REGION Network 156
   RUNG wire#powerrail
      Move(in := "Carrier_57_SDCFaultCode", out1 => "DB_SDC_EMS_TA".EMS[57].TA[1].FAULT)
      wire#w1
      Move(in := "Carrier_57_SDCFaultCode", out1 => "EMS".Carrier[57].SDC_IN.CarrierDriveFaults)
   END_RUNG
   RUNG wire#powerrail
      Contact( "IndiconTempDebugON" )
   END_RUNG wire#w1
   // the same network as SCL:
   "DB_SDC_EMS_TA".EMS[57].TA[1].FAULT := "Carrier_57_SDCFaultCode";
   IF TRUE OR "IndiconTempDebugON" THEN
       "EMS".Carrier[57].SDC_IN.CarrierDriveFaults := "Carrier_57_SDCFaultCode";
   END_IF;
END_REGION

REGION Network 157
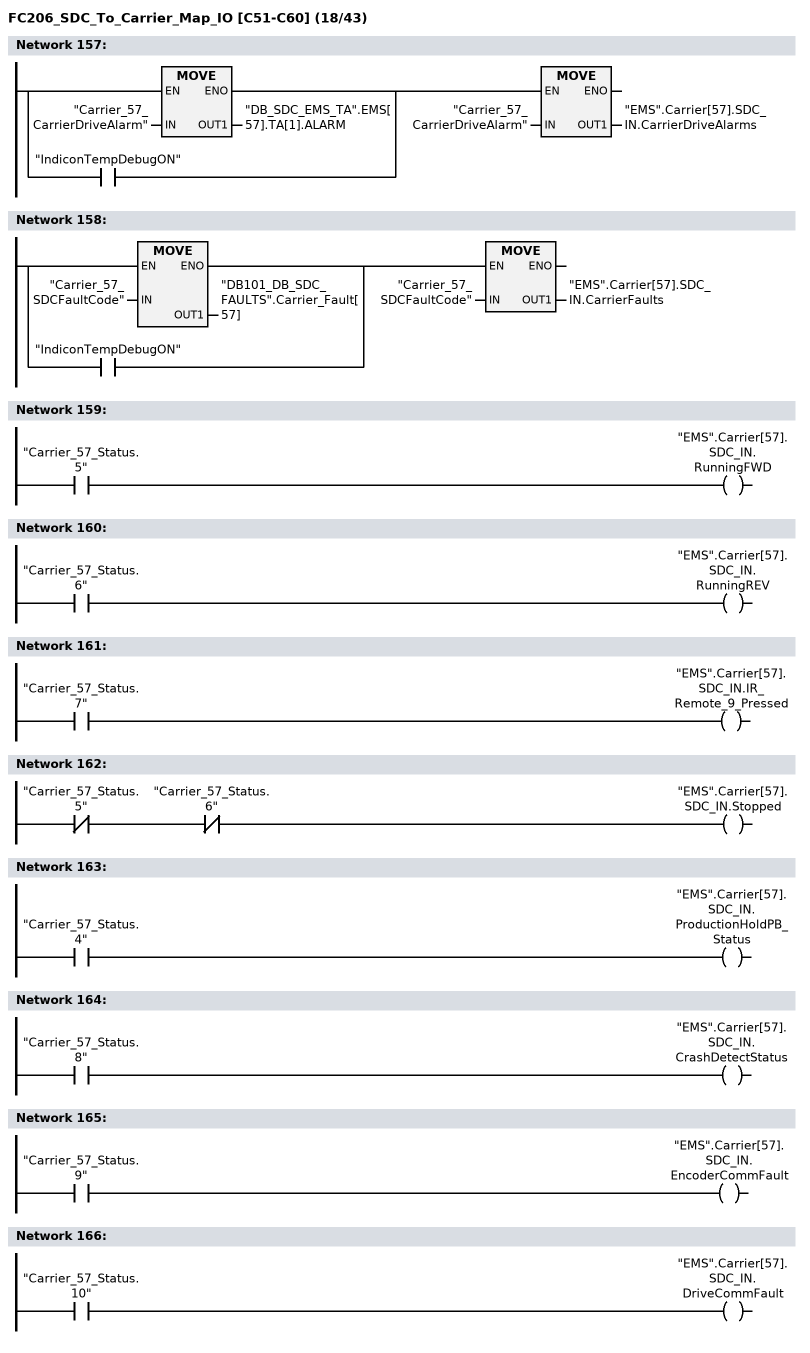
   RUNG wire#powerrail
      Move(in := "Carrier_57_CarrierDriveAlarm", out1 => "DB_SDC_EMS_TA".EMS[57].TA[1].ALARM)
      wire#w1
      Move(in := "Carrier_57_CarrierDriveAlarm", out1 => "EMS".Carrier[57].SDC_IN.CarrierDriveAlarms)
   END_RUNG
   RUNG wire#powerrail
      Contact( "IndiconTempDebugON" )
   END_RUNG wire#w1
   // the same network as SCL:
   "DB_SDC_EMS_TA".EMS[57].TA[1].ALARM := "Carrier_57_CarrierDriveAlarm";
   IF TRUE OR "IndiconTempDebugON" THEN
       "EMS".Carrier[57].SDC_IN.CarrierDriveAlarms := "Carrier_57_CarrierDriveAlarm";
   END_IF;
END_REGION

REGION Network 158
   RUNG wire#powerrail
      Move(in := "Carrier_57_SDCFaultCode", out1 => "DB101_DB_SDC_FAULTS".Carrier_Fault[57])
      wire#w1
      Move(in := "Carrier_57_SDCFaultCode", out1 => "EMS".Carrier[57].SDC_IN.CarrierFaults)
   END_RUNG
   RUNG wire#powerrail
      Contact( "IndiconTempDebugON" )
   END_RUNG wire#w1
   // the same network as SCL:
   "DB101_DB_SDC_FAULTS".Carrier_Fault[57] := "Carrier_57_SDCFaultCode";
   IF TRUE OR "IndiconTempDebugON" THEN
       "EMS".Carrier[57].SDC_IN.CarrierFaults := "Carrier_57_SDCFaultCode";
   END_IF;
END_REGION

REGION Network 159
   RUNG wire#powerrail
      Contact( "Carrier_57_Status.5" )
      Coil( "EMS".Carrier[57].SDC_IN.RunningFWD )
   END_RUNG
   // the same network as SCL:
   "EMS".Carrier[57].SDC_IN.RunningFWD := "Carrier_57_Status.5";
END_REGION

REGION Network 160
   RUNG wire#powerrail
      Contact( "Carrier_57_Status.6" )
      Coil( "EMS".Carrier[57].SDC_IN.RunningREV )
   END_RUNG
   // the same network as SCL:
   "EMS".Carrier[57].SDC_IN.RunningREV := "Carrier_57_Status.6";
END_REGION

REGION Network 161
   RUNG wire#powerrail
      Contact( "Carrier_57_Status.7" )
      Coil( "EMS".Carrier[57].SDC_IN.IR_Remote_9_Pressed )
   END_RUNG
   // the same network as SCL:
   "EMS".Carrier[57].SDC_IN.IR_Remote_9_Pressed := "Carrier_57_Status.7";
END_REGION

REGION Network 162
   RUNG wire#powerrail
      I_Contact( "Carrier_57_Status.5" )
      I_Contact( "Carrier_57_Status.6" )
      Coil( "EMS".Carrier[57].SDC_IN.Stopped )
   END_RUNG
   // the same network as SCL:
   "EMS".Carrier[57].SDC_IN.Stopped := NOT "Carrier_57_Status.5" AND NOT "Carrier_57_Status.6";
END_REGION

REGION Network 163
   RUNG wire#powerrail
      Contact( "Carrier_57_Status.4" )
      Coil( "EMS".Carrier[57].SDC_IN.ProductionHoldPB_Status )
   END_RUNG
   // the same network as SCL:
   "EMS".Carrier[57].SDC_IN.ProductionHoldPB_Status := "Carrier_57_Status.4";
END_REGION

REGION Network 164
   RUNG wire#powerrail
      Contact( "Carrier_57_Status.8" )
      Coil( "EMS".Carrier[57].SDC_IN.CrashDetectStatus )
   END_RUNG
   // the same network as SCL:
   "EMS".Carrier[57].SDC_IN.CrashDetectStatus := "Carrier_57_Status.8";
END_REGION

REGION Network 165
   RUNG wire#powerrail
      Contact( "Carrier_57_Status.9" )
      Coil( "EMS".Carrier[57].SDC_IN.EncoderCommFault )
   END_RUNG
   // the same network as SCL:
   "EMS".Carrier[57].SDC_IN.EncoderCommFault := "Carrier_57_Status.9";
END_REGION

REGION Network 166
   RUNG wire#powerrail
      Contact( "Carrier_57_Status.10" )
      Coil( "EMS".Carrier[57].SDC_IN.DriveCommFault )
   END_RUNG
   // the same network as SCL:
   "EMS".Carrier[57].SDC_IN.DriveCommFault := "Carrier_57_Status.10";
END_REGION

REGION Network 167
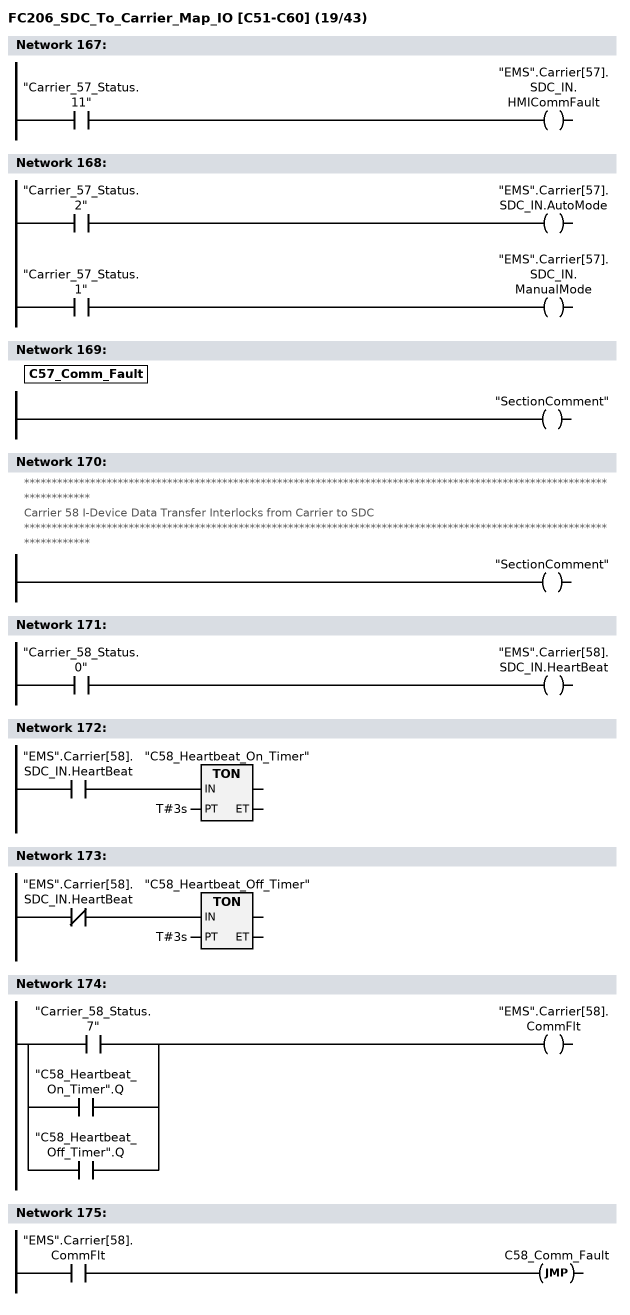
   RUNG wire#powerrail
      Contact( "Carrier_57_Status.11" )
      Coil( "EMS".Carrier[57].SDC_IN.HMICommFault )
   END_RUNG
   // the same network as SCL:
   "EMS".Carrier[57].SDC_IN.HMICommFault := "Carrier_57_Status.11";
END_REGION

REGION Network 168
   RUNG wire#powerrail
      Contact( "Carrier_57_Status.2" )
      Coil( "EMS".Carrier[57].SDC_IN.AutoMode )
   END_RUNG
   RUNG wire#powerrail
      Contact( "Carrier_57_Status.1" )
      Coil( "EMS".Carrier[57].SDC_IN.ManualMode )
   END_RUNG
   // the same network as SCL:
   "EMS".Carrier[57].SDC_IN.AutoMode := "Carrier_57_Status.2";
   "EMS".Carrier[57].SDC_IN.ManualMode := "Carrier_57_Status.1";
END_REGION

REGION Network 169
   Label( C57_Comm_Fault )
   RUNG wire#powerrail
      Coil( "SectionComment" )
   END_RUNG
   // the same network as SCL:
   C57_Comm_Fault:
   "SectionComment" := TRUE;
END_REGION

REGION Network 170
   // **********************************************************************************************************************
   // 
   // Carrier 58 I-Device Data Transfer Interlocks from Carrier to SDC
   // 
   // **********************************************************************************************************************
   RUNG wire#powerrail
      Coil( "SectionComment" )
   END_RUNG
   // the same network as SCL:
   "SectionComment" := TRUE;
END_REGION

REGION Network 171
   RUNG wire#powerrail
      Contact( "Carrier_58_Status.0" )
      Coil( "EMS".Carrier[58].SDC_IN.HeartBeat )
   END_RUNG
   // the same network as SCL:
   "EMS".Carrier[58].SDC_IN.HeartBeat := "Carrier_58_Status.0";
END_REGION

REGION Network 172
   "C58_Heartbeat_On_Timer".TON(IN := "EMS".Carrier[58].SDC_IN.HeartBeat, PT := T#3s);
END_REGION

REGION Network 173
   "C58_Heartbeat_Off_Timer".TON(IN := NOT "EMS".Carrier[58].SDC_IN.HeartBeat, PT := T#3s);
END_REGION

REGION Network 174
   RUNG wire#powerrail
      Contact( "Carrier_58_Status.7" )
      wire#w1
      Coil( "EMS".Carrier[58].CommFlt )
   END_RUNG
   RUNG wire#powerrail
      Contact( "C58_Heartbeat_On_Timer".Q )
   END_RUNG wire#w1
   RUNG wire#powerrail
      Contact( "C58_Heartbeat_Off_Timer".Q )
   END_RUNG wire#w1
   // the same network as SCL:
   "EMS".Carrier[58].CommFlt := "Carrier_58_Status.7" OR "C58_Heartbeat_On_Timer".Q OR "C58_Heartbeat_Off_Timer".Q;
END_REGION

REGION Network 175
   RUNG wire#powerrail
      Contact( "EMS".Carrier[58].CommFlt )
      JumpCoil( C58_Comm_Fault )
   END_RUNG
   // the same network as SCL:
   IF "EMS".Carrier[58].CommFlt THEN GOTO C58_Comm_Fault; END_IF;
END_REGION

REGION Network 176
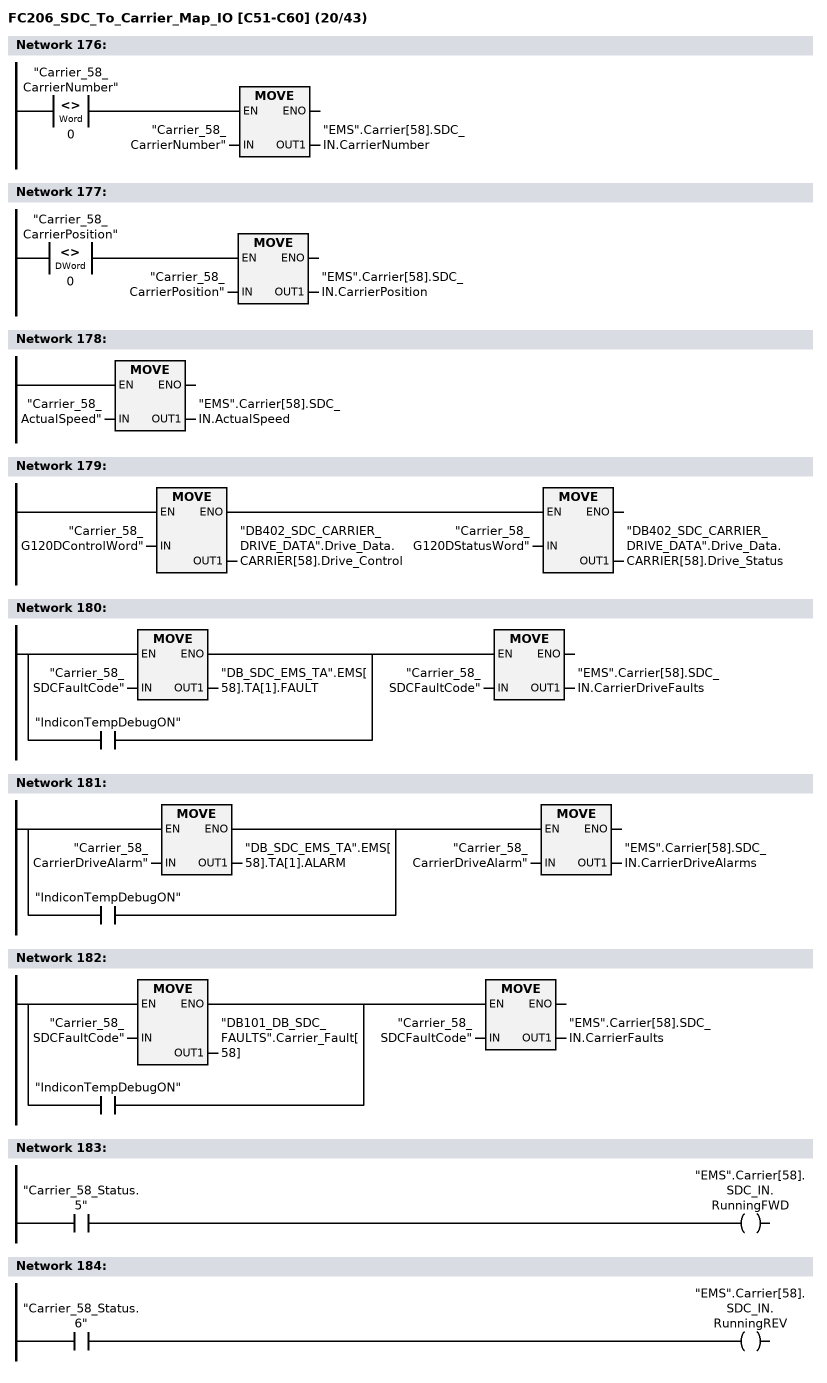
   RUNG wire#powerrail
      { S7_Templates := "SrcType := Word" } NE_Contact(in1 := "Carrier_58_CarrierNumber", in2 := 0)
      Move(in := "Carrier_58_CarrierNumber", out1 => "EMS".Carrier[58].SDC_IN.CarrierNumber)
   END_RUNG
   // the same network as SCL:
   IF "Carrier_58_CarrierNumber" <> 0 THEN
       "EMS".Carrier[58].SDC_IN.CarrierNumber := "Carrier_58_CarrierNumber";
   END_IF;
END_REGION

REGION Network 177
   RUNG wire#powerrail
      { S7_Templates := "SrcType := DWord" } NE_Contact(in1 := "Carrier_58_CarrierPosition", in2 := 0)
      Move(in := "Carrier_58_CarrierPosition", out1 => "EMS".Carrier[58].SDC_IN.CarrierPosition)
   END_RUNG
   // the same network as SCL:
   IF "Carrier_58_CarrierPosition" <> 0 THEN
       "EMS".Carrier[58].SDC_IN.CarrierPosition := "Carrier_58_CarrierPosition";
   END_IF;
END_REGION

REGION Network 178
   RUNG wire#powerrail
      Move(in := "Carrier_58_ActualSpeed", out1 => "EMS".Carrier[58].SDC_IN.ActualSpeed)
   END_RUNG
   // the same network as SCL:
   "EMS".Carrier[58].SDC_IN.ActualSpeed := "Carrier_58_ActualSpeed";
END_REGION

REGION Network 179
   RUNG wire#powerrail
      Move(in := "Carrier_58_G120DControlWord", out1 => "DB402_SDC_CARRIER_DRIVE_DATA".Drive_Data.CARRIER[58].Drive_Control)
      Move(in := "Carrier_58_G120DStatusWord", out1 => "DB402_SDC_CARRIER_DRIVE_DATA".Drive_Data.CARRIER[58].Drive_Status)
   END_RUNG
   // the same network as SCL:
   "DB402_SDC_CARRIER_DRIVE_DATA".Drive_Data.CARRIER[58].Drive_Control := "Carrier_58_G120DControlWord";
   "DB402_SDC_CARRIER_DRIVE_DATA".Drive_Data.CARRIER[58].Drive_Status := "Carrier_58_G120DStatusWord";
END_REGION

REGION Network 180
   RUNG wire#powerrail
      Move(in := "Carrier_58_SDCFaultCode", out1 => "DB_SDC_EMS_TA".EMS[58].TA[1].FAULT)
      wire#w1
      Move(in := "Carrier_58_SDCFaultCode", out1 => "EMS".Carrier[58].SDC_IN.CarrierDriveFaults)
   END_RUNG
   RUNG wire#powerrail
      Contact( "IndiconTempDebugON" )
   END_RUNG wire#w1
   // the same network as SCL:
   "DB_SDC_EMS_TA".EMS[58].TA[1].FAULT := "Carrier_58_SDCFaultCode";
   IF TRUE OR "IndiconTempDebugON" THEN
       "EMS".Carrier[58].SDC_IN.CarrierDriveFaults := "Carrier_58_SDCFaultCode";
   END_IF;
END_REGION

REGION Network 181
   RUNG wire#powerrail
      Move(in := "Carrier_58_CarrierDriveAlarm", out1 => "DB_SDC_EMS_TA".EMS[58].TA[1].ALARM)
      wire#w1
      Move(in := "Carrier_58_CarrierDriveAlarm", out1 => "EMS".Carrier[58].SDC_IN.CarrierDriveAlarms)
   END_RUNG
   RUNG wire#powerrail
      Contact( "IndiconTempDebugON" )
   END_RUNG wire#w1
   // the same network as SCL:
   "DB_SDC_EMS_TA".EMS[58].TA[1].ALARM := "Carrier_58_CarrierDriveAlarm";
   IF TRUE OR "IndiconTempDebugON" THEN
       "EMS".Carrier[58].SDC_IN.CarrierDriveAlarms := "Carrier_58_CarrierDriveAlarm";
   END_IF;
END_REGION

REGION Network 182
   RUNG wire#powerrail
      Move(in := "Carrier_58_SDCFaultCode", out1 => "DB101_DB_SDC_FAULTS".Carrier_Fault[58])
      wire#w1
      Move(in := "Carrier_58_SDCFaultCode", out1 => "EMS".Carrier[58].SDC_IN.CarrierFaults)
   END_RUNG
   RUNG wire#powerrail
      Contact( "IndiconTempDebugON" )
   END_RUNG wire#w1
   // the same network as SCL:
   "DB101_DB_SDC_FAULTS".Carrier_Fault[58] := "Carrier_58_SDCFaultCode";
   IF TRUE OR "IndiconTempDebugON" THEN
       "EMS".Carrier[58].SDC_IN.CarrierFaults := "Carrier_58_SDCFaultCode";
   END_IF;
END_REGION

REGION Network 183
   RUNG wire#powerrail
      Contact( "Carrier_58_Status.5" )
      Coil( "EMS".Carrier[58].SDC_IN.RunningFWD )
   END_RUNG
   // the same network as SCL:
   "EMS".Carrier[58].SDC_IN.RunningFWD := "Carrier_58_Status.5";
END_REGION

REGION Network 184
   RUNG wire#powerrail
      Contact( "Carrier_58_Status.6" )
      Coil( "EMS".Carrier[58].SDC_IN.RunningREV )
   END_RUNG
   // the same network as SCL:
   "EMS".Carrier[58].SDC_IN.RunningREV := "Carrier_58_Status.6";
END_REGION

REGION Network 185
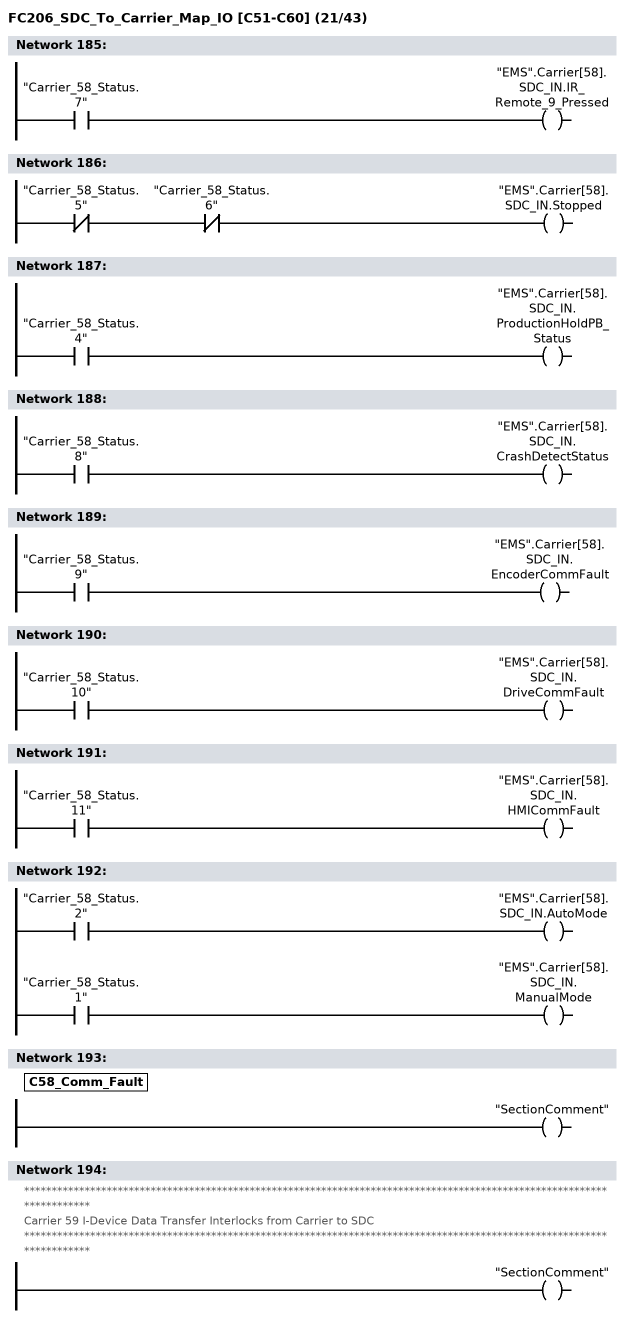
   RUNG wire#powerrail
      Contact( "Carrier_58_Status.7" )
      Coil( "EMS".Carrier[58].SDC_IN.IR_Remote_9_Pressed )
   END_RUNG
   // the same network as SCL:
   "EMS".Carrier[58].SDC_IN.IR_Remote_9_Pressed := "Carrier_58_Status.7";
END_REGION

REGION Network 186
   RUNG wire#powerrail
      I_Contact( "Carrier_58_Status.5" )
      I_Contact( "Carrier_58_Status.6" )
      Coil( "EMS".Carrier[58].SDC_IN.Stopped )
   END_RUNG
   // the same network as SCL:
   "EMS".Carrier[58].SDC_IN.Stopped := NOT "Carrier_58_Status.5" AND NOT "Carrier_58_Status.6";
END_REGION

REGION Network 187
   RUNG wire#powerrail
      Contact( "Carrier_58_Status.4" )
      Coil( "EMS".Carrier[58].SDC_IN.ProductionHoldPB_Status )
   END_RUNG
   // the same network as SCL:
   "EMS".Carrier[58].SDC_IN.ProductionHoldPB_Status := "Carrier_58_Status.4";
END_REGION

REGION Network 188
   RUNG wire#powerrail
      Contact( "Carrier_58_Status.8" )
      Coil( "EMS".Carrier[58].SDC_IN.CrashDetectStatus )
   END_RUNG
   // the same network as SCL:
   "EMS".Carrier[58].SDC_IN.CrashDetectStatus := "Carrier_58_Status.8";
END_REGION

REGION Network 189
   RUNG wire#powerrail
      Contact( "Carrier_58_Status.9" )
      Coil( "EMS".Carrier[58].SDC_IN.EncoderCommFault )
   END_RUNG
   // the same network as SCL:
   "EMS".Carrier[58].SDC_IN.EncoderCommFault := "Carrier_58_Status.9";
END_REGION

REGION Network 190
   RUNG wire#powerrail
      Contact( "Carrier_58_Status.10" )
      Coil( "EMS".Carrier[58].SDC_IN.DriveCommFault )
   END_RUNG
   // the same network as SCL:
   "EMS".Carrier[58].SDC_IN.DriveCommFault := "Carrier_58_Status.10";
END_REGION

REGION Network 191
   RUNG wire#powerrail
      Contact( "Carrier_58_Status.11" )
      Coil( "EMS".Carrier[58].SDC_IN.HMICommFault )
   END_RUNG
   // the same network as SCL:
   "EMS".Carrier[58].SDC_IN.HMICommFault := "Carrier_58_Status.11";
END_REGION

REGION Network 192
   RUNG wire#powerrail
      Contact( "Carrier_58_Status.2" )
      Coil( "EMS".Carrier[58].SDC_IN.AutoMode )
   END_RUNG
   RUNG wire#powerrail
      Contact( "Carrier_58_Status.1" )
      Coil( "EMS".Carrier[58].SDC_IN.ManualMode )
   END_RUNG
   // the same network as SCL:
   "EMS".Carrier[58].SDC_IN.AutoMode := "Carrier_58_Status.2";
   "EMS".Carrier[58].SDC_IN.ManualMode := "Carrier_58_Status.1";
END_REGION

REGION Network 193
   Label( C58_Comm_Fault )
   RUNG wire#powerrail
      Coil( "SectionComment" )
   END_RUNG
   // the same network as SCL:
   C58_Comm_Fault:
   "SectionComment" := TRUE;
END_REGION

REGION Network 194
   // **********************************************************************************************************************
   // 
   // Carrier 59 I-Device Data Transfer Interlocks from Carrier to SDC
   // 
   // **********************************************************************************************************************
   RUNG wire#powerrail
      Coil( "SectionComment" )
   END_RUNG
   // the same network as SCL:
   "SectionComment" := TRUE;
END_REGION

REGION Network 195
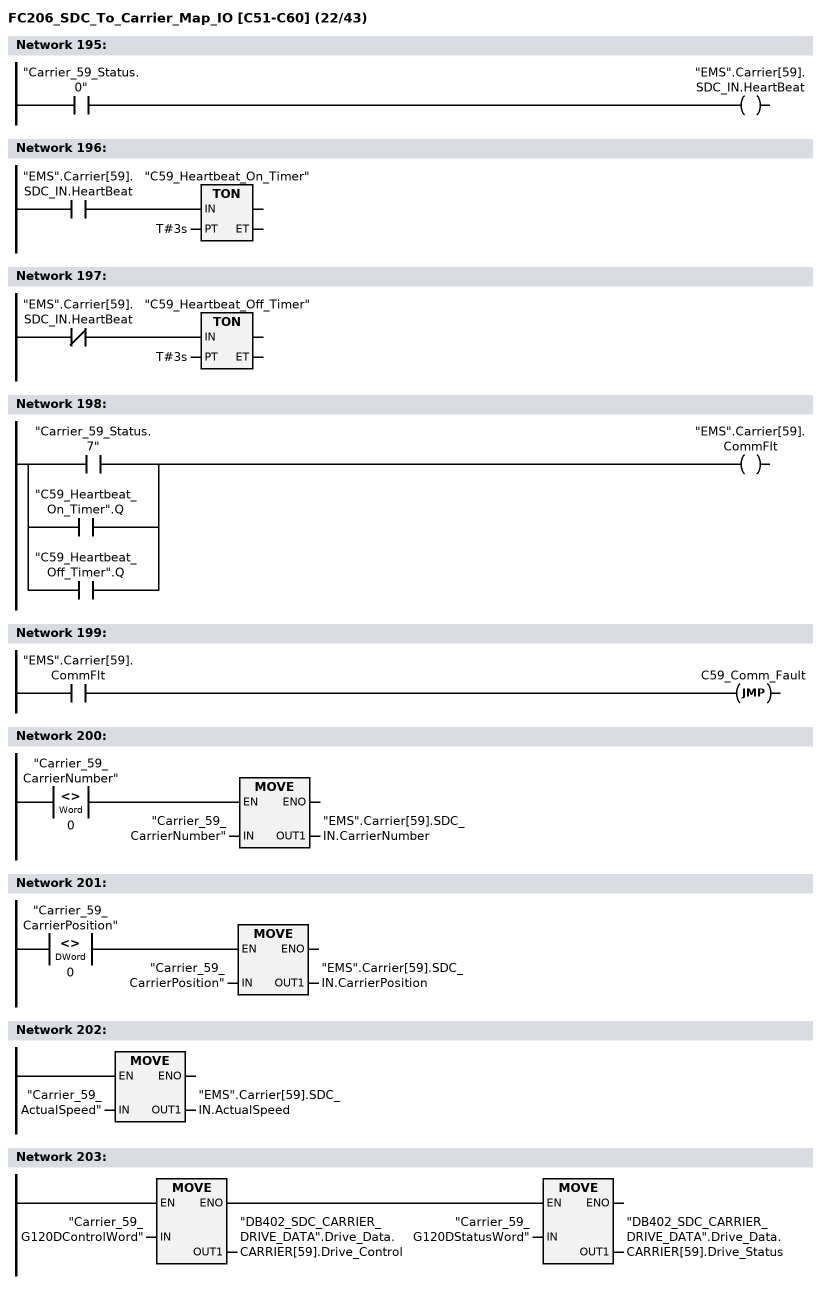
   RUNG wire#powerrail
      Contact( "Carrier_59_Status.0" )
      Coil( "EMS".Carrier[59].SDC_IN.HeartBeat )
   END_RUNG
   // the same network as SCL:
   "EMS".Carrier[59].SDC_IN.HeartBeat := "Carrier_59_Status.0";
END_REGION

REGION Network 196
   "C59_Heartbeat_On_Timer".TON(IN := "EMS".Carrier[59].SDC_IN.HeartBeat, PT := T#3s);
END_REGION

REGION Network 197
   "C59_Heartbeat_Off_Timer".TON(IN := NOT "EMS".Carrier[59].SDC_IN.HeartBeat, PT := T#3s);
END_REGION

REGION Network 198
   RUNG wire#powerrail
      Contact( "Carrier_59_Status.7" )
      wire#w1
      Coil( "EMS".Carrier[59].CommFlt )
   END_RUNG
   RUNG wire#powerrail
      Contact( "C59_Heartbeat_On_Timer".Q )
   END_RUNG wire#w1
   RUNG wire#powerrail
      Contact( "C59_Heartbeat_Off_Timer".Q )
   END_RUNG wire#w1
   // the same network as SCL:
   "EMS".Carrier[59].CommFlt := "Carrier_59_Status.7" OR "C59_Heartbeat_On_Timer".Q OR "C59_Heartbeat_Off_Timer".Q;
END_REGION

REGION Network 199
   RUNG wire#powerrail
      Contact( "EMS".Carrier[59].CommFlt )
      JumpCoil( C59_Comm_Fault )
   END_RUNG
   // the same network as SCL:
   IF "EMS".Carrier[59].CommFlt THEN GOTO C59_Comm_Fault; END_IF;
END_REGION

REGION Network 200
   RUNG wire#powerrail
      { S7_Templates := "SrcType := Word" } NE_Contact(in1 := "Carrier_59_CarrierNumber", in2 := 0)
      Move(in := "Carrier_59_CarrierNumber", out1 => "EMS".Carrier[59].SDC_IN.CarrierNumber)
   END_RUNG
   // the same network as SCL:
   IF "Carrier_59_CarrierNumber" <> 0 THEN
       "EMS".Carrier[59].SDC_IN.CarrierNumber := "Carrier_59_CarrierNumber";
   END_IF;
END_REGION

REGION Network 201
   RUNG wire#powerrail
      { S7_Templates := "SrcType := DWord" } NE_Contact(in1 := "Carrier_59_CarrierPosition", in2 := 0)
      Move(in := "Carrier_59_CarrierPosition", out1 => "EMS".Carrier[59].SDC_IN.CarrierPosition)
   END_RUNG
   // the same network as SCL:
   IF "Carrier_59_CarrierPosition" <> 0 THEN
       "EMS".Carrier[59].SDC_IN.CarrierPosition := "Carrier_59_CarrierPosition";
   END_IF;
END_REGION

REGION Network 202
   RUNG wire#powerrail
      Move(in := "Carrier_59_ActualSpeed", out1 => "EMS".Carrier[59].SDC_IN.ActualSpeed)
   END_RUNG
   // the same network as SCL:
   "EMS".Carrier[59].SDC_IN.ActualSpeed := "Carrier_59_ActualSpeed";
END_REGION

REGION Network 203
   RUNG wire#powerrail
      Move(in := "Carrier_59_G120DControlWord", out1 => "DB402_SDC_CARRIER_DRIVE_DATA".Drive_Data.CARRIER[59].Drive_Control)
      Move(in := "Carrier_59_G120DStatusWord", out1 => "DB402_SDC_CARRIER_DRIVE_DATA".Drive_Data.CARRIER[59].Drive_Status)
   END_RUNG
   // the same network as SCL:
   "DB402_SDC_CARRIER_DRIVE_DATA".Drive_Data.CARRIER[59].Drive_Control := "Carrier_59_G120DControlWord";
   "DB402_SDC_CARRIER_DRIVE_DATA".Drive_Data.CARRIER[59].Drive_Status := "Carrier_59_G120DStatusWord";
END_REGION

REGION Network 204
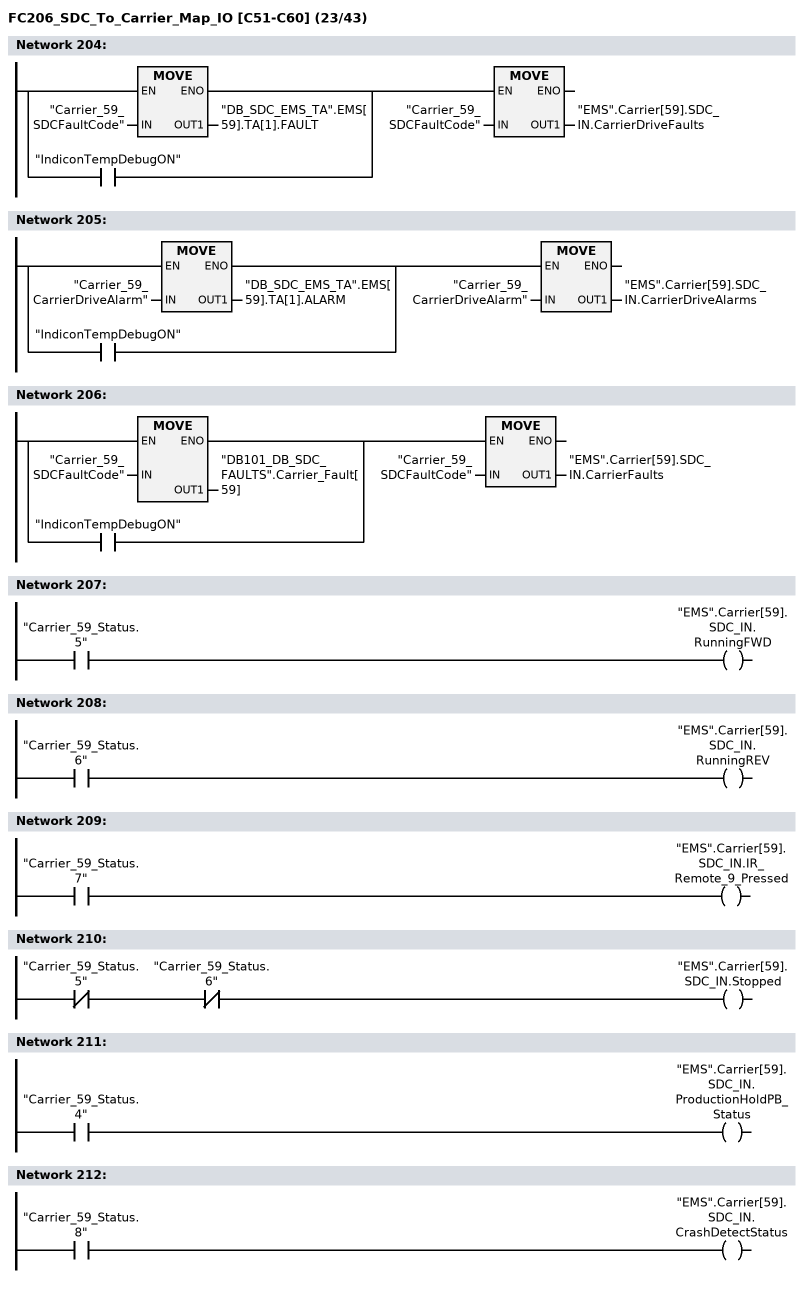
   RUNG wire#powerrail
      Move(in := "Carrier_59_SDCFaultCode", out1 => "DB_SDC_EMS_TA".EMS[59].TA[1].FAULT)
      wire#w1
      Move(in := "Carrier_59_SDCFaultCode", out1 => "EMS".Carrier[59].SDC_IN.CarrierDriveFaults)
   END_RUNG
   RUNG wire#powerrail
      Contact( "IndiconTempDebugON" )
   END_RUNG wire#w1
   // the same network as SCL:
   "DB_SDC_EMS_TA".EMS[59].TA[1].FAULT := "Carrier_59_SDCFaultCode";
   IF TRUE OR "IndiconTempDebugON" THEN
       "EMS".Carrier[59].SDC_IN.CarrierDriveFaults := "Carrier_59_SDCFaultCode";
   END_IF;
END_REGION

REGION Network 205
   RUNG wire#powerrail
      Move(in := "Carrier_59_CarrierDriveAlarm", out1 => "DB_SDC_EMS_TA".EMS[59].TA[1].ALARM)
      wire#w1
      Move(in := "Carrier_59_CarrierDriveAlarm", out1 => "EMS".Carrier[59].SDC_IN.CarrierDriveAlarms)
   END_RUNG
   RUNG wire#powerrail
      Contact( "IndiconTempDebugON" )
   END_RUNG wire#w1
   // the same network as SCL:
   "DB_SDC_EMS_TA".EMS[59].TA[1].ALARM := "Carrier_59_CarrierDriveAlarm";
   IF TRUE OR "IndiconTempDebugON" THEN
       "EMS".Carrier[59].SDC_IN.CarrierDriveAlarms := "Carrier_59_CarrierDriveAlarm";
   END_IF;
END_REGION

REGION Network 206
   RUNG wire#powerrail
      Move(in := "Carrier_59_SDCFaultCode", out1 => "DB101_DB_SDC_FAULTS".Carrier_Fault[59])
      wire#w1
      Move(in := "Carrier_59_SDCFaultCode", out1 => "EMS".Carrier[59].SDC_IN.CarrierFaults)
   END_RUNG
   RUNG wire#powerrail
      Contact( "IndiconTempDebugON" )
   END_RUNG wire#w1
   // the same network as SCL:
   "DB101_DB_SDC_FAULTS".Carrier_Fault[59] := "Carrier_59_SDCFaultCode";
   IF TRUE OR "IndiconTempDebugON" THEN
       "EMS".Carrier[59].SDC_IN.CarrierFaults := "Carrier_59_SDCFaultCode";
   END_IF;
END_REGION

REGION Network 207
   RUNG wire#powerrail
      Contact( "Carrier_59_Status.5" )
      Coil( "EMS".Carrier[59].SDC_IN.RunningFWD )
   END_RUNG
   // the same network as SCL:
   "EMS".Carrier[59].SDC_IN.RunningFWD := "Carrier_59_Status.5";
END_REGION

REGION Network 208
   RUNG wire#powerrail
      Contact( "Carrier_59_Status.6" )
      Coil( "EMS".Carrier[59].SDC_IN.RunningREV )
   END_RUNG
   // the same network as SCL:
   "EMS".Carrier[59].SDC_IN.RunningREV := "Carrier_59_Status.6";
END_REGION

REGION Network 209
   RUNG wire#powerrail
      Contact( "Carrier_59_Status.7" )
      Coil( "EMS".Carrier[59].SDC_IN.IR_Remote_9_Pressed )
   END_RUNG
   // the same network as SCL:
   "EMS".Carrier[59].SDC_IN.IR_Remote_9_Pressed := "Carrier_59_Status.7";
END_REGION

REGION Network 210
   RUNG wire#powerrail
      I_Contact( "Carrier_59_Status.5" )
      I_Contact( "Carrier_59_Status.6" )
      Coil( "EMS".Carrier[59].SDC_IN.Stopped )
   END_RUNG
   // the same network as SCL:
   "EMS".Carrier[59].SDC_IN.Stopped := NOT "Carrier_59_Status.5" AND NOT "Carrier_59_Status.6";
END_REGION

REGION Network 211
   RUNG wire#powerrail
      Contact( "Carrier_59_Status.4" )
      Coil( "EMS".Carrier[59].SDC_IN.ProductionHoldPB_Status )
   END_RUNG
   // the same network as SCL:
   "EMS".Carrier[59].SDC_IN.ProductionHoldPB_Status := "Carrier_59_Status.4";
END_REGION

REGION Network 212
   RUNG wire#powerrail
      Contact( "Carrier_59_Status.8" )
      Coil( "EMS".Carrier[59].SDC_IN.CrashDetectStatus )
   END_RUNG
   // the same network as SCL:
   "EMS".Carrier[59].SDC_IN.CrashDetectStatus := "Carrier_59_Status.8";
END_REGION

REGION Network 213
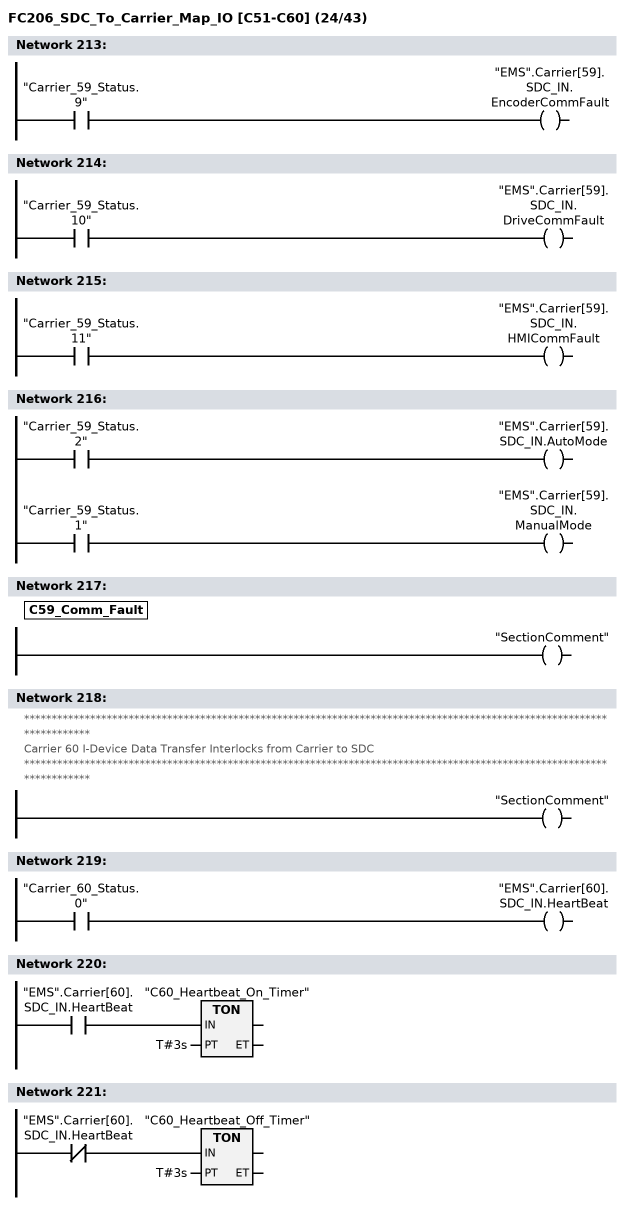
   RUNG wire#powerrail
      Contact( "Carrier_59_Status.9" )
      Coil( "EMS".Carrier[59].SDC_IN.EncoderCommFault )
   END_RUNG
   // the same network as SCL:
   "EMS".Carrier[59].SDC_IN.EncoderCommFault := "Carrier_59_Status.9";
END_REGION

REGION Network 214
   RUNG wire#powerrail
      Contact( "Carrier_59_Status.10" )
      Coil( "EMS".Carrier[59].SDC_IN.DriveCommFault )
   END_RUNG
   // the same network as SCL:
   "EMS".Carrier[59].SDC_IN.DriveCommFault := "Carrier_59_Status.10";
END_REGION

REGION Network 215
   RUNG wire#powerrail
      Contact( "Carrier_59_Status.11" )
      Coil( "EMS".Carrier[59].SDC_IN.HMICommFault )
   END_RUNG
   // the same network as SCL:
   "EMS".Carrier[59].SDC_IN.HMICommFault := "Carrier_59_Status.11";
END_REGION

REGION Network 216
   RUNG wire#powerrail
      Contact( "Carrier_59_Status.2" )
      Coil( "EMS".Carrier[59].SDC_IN.AutoMode )
   END_RUNG
   RUNG wire#powerrail
      Contact( "Carrier_59_Status.1" )
      Coil( "EMS".Carrier[59].SDC_IN.ManualMode )
   END_RUNG
   // the same network as SCL:
   "EMS".Carrier[59].SDC_IN.AutoMode := "Carrier_59_Status.2";
   "EMS".Carrier[59].SDC_IN.ManualMode := "Carrier_59_Status.1";
END_REGION

REGION Network 217
   Label( C59_Comm_Fault )
   RUNG wire#powerrail
      Coil( "SectionComment" )
   END_RUNG
   // the same network as SCL:
   C59_Comm_Fault:
   "SectionComment" := TRUE;
END_REGION

REGION Network 218
   // **********************************************************************************************************************
   // 
   // Carrier 60 I-Device Data Transfer Interlocks from Carrier to SDC
   // 
   // **********************************************************************************************************************
   RUNG wire#powerrail
      Coil( "SectionComment" )
   END_RUNG
   // the same network as SCL:
   "SectionComment" := TRUE;
END_REGION

REGION Network 219
   RUNG wire#powerrail
      Contact( "Carrier_60_Status.0" )
      Coil( "EMS".Carrier[60].SDC_IN.HeartBeat )
   END_RUNG
   // the same network as SCL:
   "EMS".Carrier[60].SDC_IN.HeartBeat := "Carrier_60_Status.0";
END_REGION

REGION Network 220
   "C60_Heartbeat_On_Timer".TON(IN := "EMS".Carrier[60].SDC_IN.HeartBeat, PT := T#3s);
END_REGION

REGION Network 221
   "C60_Heartbeat_Off_Timer".TON(IN := NOT "EMS".Carrier[60].SDC_IN.HeartBeat, PT := T#3s);
END_REGION

REGION Network 222
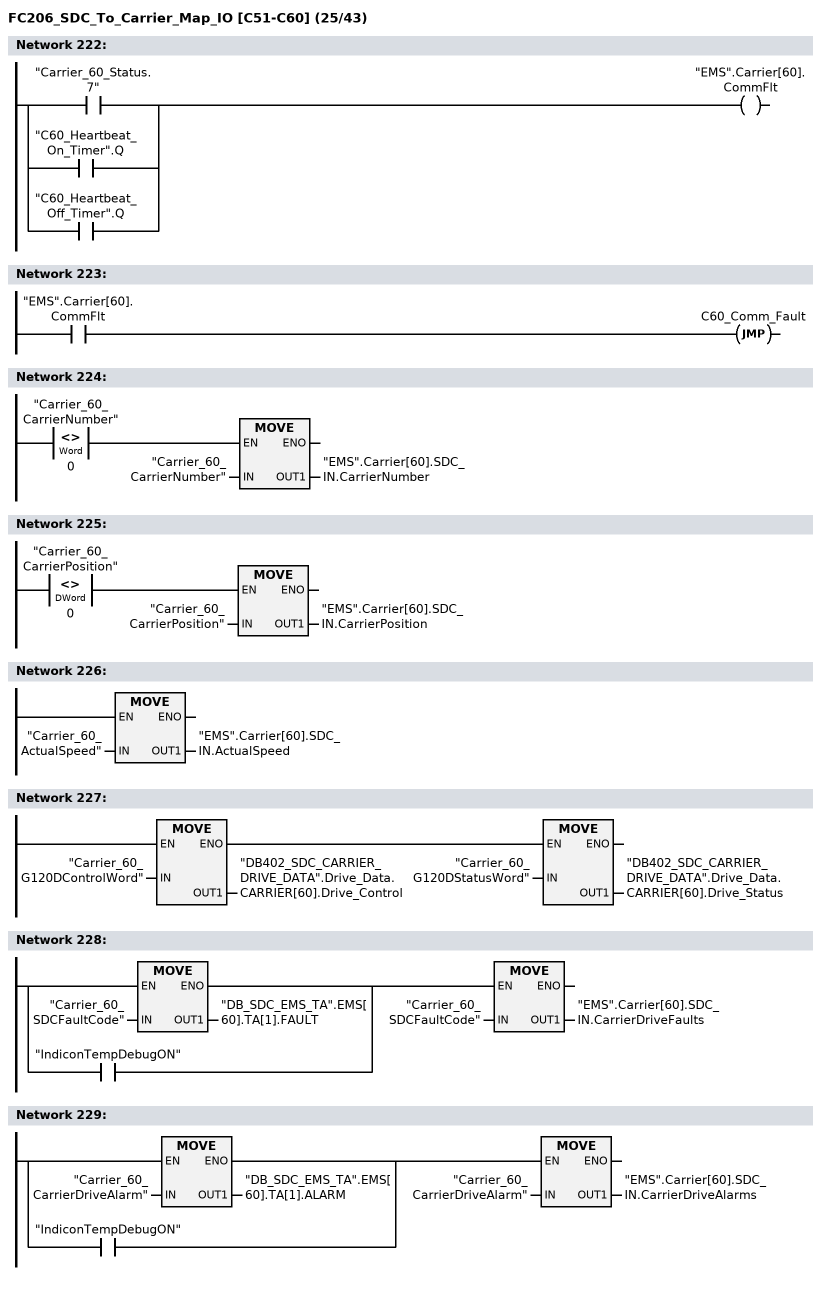
   RUNG wire#powerrail
      Contact( "Carrier_60_Status.7" )
      wire#w1
      Coil( "EMS".Carrier[60].CommFlt )
   END_RUNG
   RUNG wire#powerrail
      Contact( "C60_Heartbeat_On_Timer".Q )
   END_RUNG wire#w1
   RUNG wire#powerrail
      Contact( "C60_Heartbeat_Off_Timer".Q )
   END_RUNG wire#w1
   // the same network as SCL:
   "EMS".Carrier[60].CommFlt := "Carrier_60_Status.7" OR "C60_Heartbeat_On_Timer".Q OR "C60_Heartbeat_Off_Timer".Q;
END_REGION

REGION Network 223
   RUNG wire#powerrail
      Contact( "EMS".Carrier[60].CommFlt )
      JumpCoil( C60_Comm_Fault )
   END_RUNG
   // the same network as SCL:
   IF "EMS".Carrier[60].CommFlt THEN GOTO C60_Comm_Fault; END_IF;
END_REGION

REGION Network 224
   RUNG wire#powerrail
      { S7_Templates := "SrcType := Word" } NE_Contact(in1 := "Carrier_60_CarrierNumber", in2 := 0)
      Move(in := "Carrier_60_CarrierNumber", out1 => "EMS".Carrier[60].SDC_IN.CarrierNumber)
   END_RUNG
   // the same network as SCL:
   IF "Carrier_60_CarrierNumber" <> 0 THEN
       "EMS".Carrier[60].SDC_IN.CarrierNumber := "Carrier_60_CarrierNumber";
   END_IF;
END_REGION

REGION Network 225
   RUNG wire#powerrail
      { S7_Templates := "SrcType := DWord" } NE_Contact(in1 := "Carrier_60_CarrierPosition", in2 := 0)
      Move(in := "Carrier_60_CarrierPosition", out1 => "EMS".Carrier[60].SDC_IN.CarrierPosition)
   END_RUNG
   // the same network as SCL:
   IF "Carrier_60_CarrierPosition" <> 0 THEN
       "EMS".Carrier[60].SDC_IN.CarrierPosition := "Carrier_60_CarrierPosition";
   END_IF;
END_REGION

REGION Network 226
   RUNG wire#powerrail
      Move(in := "Carrier_60_ActualSpeed", out1 => "EMS".Carrier[60].SDC_IN.ActualSpeed)
   END_RUNG
   // the same network as SCL:
   "EMS".Carrier[60].SDC_IN.ActualSpeed := "Carrier_60_ActualSpeed";
END_REGION

REGION Network 227
   RUNG wire#powerrail
      Move(in := "Carrier_60_G120DControlWord", out1 => "DB402_SDC_CARRIER_DRIVE_DATA".Drive_Data.CARRIER[60].Drive_Control)
      Move(in := "Carrier_60_G120DStatusWord", out1 => "DB402_SDC_CARRIER_DRIVE_DATA".Drive_Data.CARRIER[60].Drive_Status)
   END_RUNG
   // the same network as SCL:
   "DB402_SDC_CARRIER_DRIVE_DATA".Drive_Data.CARRIER[60].Drive_Control := "Carrier_60_G120DControlWord";
   "DB402_SDC_CARRIER_DRIVE_DATA".Drive_Data.CARRIER[60].Drive_Status := "Carrier_60_G120DStatusWord";
END_REGION

REGION Network 228
   RUNG wire#powerrail
      Move(in := "Carrier_60_SDCFaultCode", out1 => "DB_SDC_EMS_TA".EMS[60].TA[1].FAULT)
      wire#w1
      Move(in := "Carrier_60_SDCFaultCode", out1 => "EMS".Carrier[60].SDC_IN.CarrierDriveFaults)
   END_RUNG
   RUNG wire#powerrail
      Contact( "IndiconTempDebugON" )
   END_RUNG wire#w1
   // the same network as SCL:
   "DB_SDC_EMS_TA".EMS[60].TA[1].FAULT := "Carrier_60_SDCFaultCode";
   IF TRUE OR "IndiconTempDebugON" THEN
       "EMS".Carrier[60].SDC_IN.CarrierDriveFaults := "Carrier_60_SDCFaultCode";
   END_IF;
END_REGION

REGION Network 229
   RUNG wire#powerrail
      Move(in := "Carrier_60_CarrierDriveAlarm", out1 => "DB_SDC_EMS_TA".EMS[60].TA[1].ALARM)
      wire#w1
      Move(in := "Carrier_60_CarrierDriveAlarm", out1 => "EMS".Carrier[60].SDC_IN.CarrierDriveAlarms)
   END_RUNG
   RUNG wire#powerrail
      Contact( "IndiconTempDebugON" )
   END_RUNG wire#w1
   // the same network as SCL:
   "DB_SDC_EMS_TA".EMS[60].TA[1].ALARM := "Carrier_60_CarrierDriveAlarm";
   IF TRUE OR "IndiconTempDebugON" THEN
       "EMS".Carrier[60].SDC_IN.CarrierDriveAlarms := "Carrier_60_CarrierDriveAlarm";
   END_IF;
END_REGION

REGION Network 230
